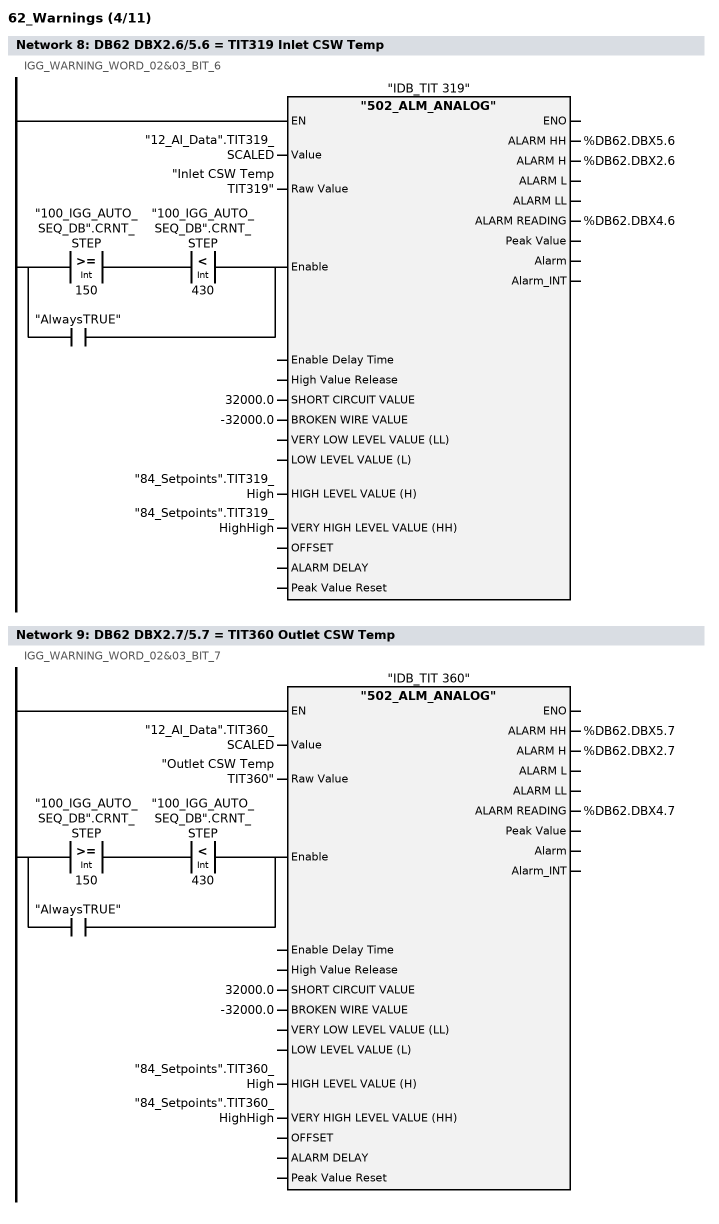
   RUNG wire#powerrail
      "IDB_TIT 319"(Enable := wire#w1, Value := "12_AI_Data".TIT319_SCALED, "Raw Value" := "Inlet CSW Temp TIT319", "SHORT CIRCUIT VALUE" := 32000.0, "BROKEN WIRE VALUE" := -32000.0, "VERY LOW LEVEL VALUE (LL)" :=, "LOW LEVEL VALUE (L)" :=, "HIGH LEVEL VALUE (H)" := "84_Setpoints".TIT319_High, "VERY HIGH LEVEL VALUE (HH)" := "84_Setpoints".TIT319_HighHigh, OFFSET :=, "ALARM DELAY" :=, "Peak Value Reset" :=, "ALARM HH" => %DB62.DBX5.6, "ALARM H" => %DB62.DBX2.6, "ALARM L" =>, "ALARM LL" =>, "ALARM READING" => %DB62.DBX4.6, "Peak Value" =>, Alarm =>, Alarm_INT =>, "Enable Delay Time" :=, "High Value Release" :=)
   END_RUNG
   RUNG wire#powerrail
      { S7_Templates := "SrcType := Int" } GE_Contact(in1 := "100_IGG_AUTO_SEQ_DB".CRNT_STEP, in2 := 150)
      { S7_Templates := "SrcType := Int" } LT_Contact(in1 := "100_IGG_AUTO_SEQ_DB".CRNT_STEP, in2 := 430)
   END_RUNG wire#w1
   RUNG wire#powerrail
      Contact( "AlwaysTRUE" )
   END_RUNG wire#w1
   // the same network as SCL:
   "IDB_TIT 319"(Value := "12_AI_Data".TIT319_SCALED,   // "502_ALM_ANALOG"
                 "Raw Value" := "Inlet CSW Temp TIT319",
                 Enable := (("100_IGG_AUTO_SEQ_DB".CRNT_STEP >= 150) AND ("100_IGG_AUTO_SEQ_DB".CRNT_STEP < 430)) OR "AlwaysTRUE",
                 "SHORT CIRCUIT VALUE" := 32000.0,
                 "BROKEN WIRE VALUE" := -32000.0,
                 "HIGH LEVEL VALUE (H)" := "84_Setpoints".TIT319_High,
                 "VERY HIGH LEVEL VALUE (HH)" := "84_Setpoints".TIT319_HighHigh,
                 "ALARM HH" => %DB62.DBX5.6,
                 "ALARM H" => %DB62.DBX2.6,
                 "ALARM READING" => %DB62.DBX4.6);
END_REGION

REGION Network 9: DB62 DBX2.7/5.7 = TIT360 Outlet CSW Temp
   // IGG_WARNING_WORD_02&03_BIT_7
   RUNG wire#powerrail
      "IDB_TIT 360"(Enable := wire#w1, Value := "12_AI_Data".TIT360_SCALED, "Raw Value" := "Outlet CSW Temp TIT360", "SHORT CIRCUIT VALUE" := 32000.0, "BROKEN WIRE VALUE" := -32000.0, "VERY LOW LEVEL VALUE (LL)" :=, "LOW LEVEL VALUE (L)" :=, "HIGH LEVEL VALUE (H)" := "84_Setpoints".TIT360_High, "VERY HIGH LEVEL VALUE (HH)" := "84_Setpoints".TIT360_HighHigh, OFFSET :=, "ALARM DELAY" :=, "Peak Value Reset" :=, "ALARM HH" => %DB62.DBX5.7, "ALARM H" => %DB62.DBX2.7, "ALARM L" =>, "ALARM LL" =>, "ALARM READING" => %DB62.DBX4.7, "Peak Value" =>, Alarm =>, Alarm_INT =>, "Enable Delay Time" :=, "High Value Release" :=)
   END_RUNG
   RUNG wire#powerrail
      { S7_Templates := "SrcType := Int" } GE_Contact(in1 := "100_IGG_AUTO_SEQ_DB".CRNT_STEP, in2 := 150)
      { S7_Templates := "SrcType := Int" } LT_Contact(in1 := "100_IGG_AUTO_SEQ_DB".CRNT_STEP, in2 := 430)
   END_RUNG wire#w1
   RUNG wire#powerrail
      Contact( "AlwaysTRUE" )
   END_RUNG wire#w1
   // the same network as SCL:
   "IDB_TIT 360"(Value := "12_AI_Data".TIT360_SCALED,   // "502_ALM_ANALOG"
                 "Raw Value" := "Outlet CSW Temp TIT360",
                 Enable := (("100_IGG_AUTO_SEQ_DB".CRNT_STEP >= 150) AND ("100_IGG_AUTO_SEQ_DB".CRNT_STEP < 430)) OR "AlwaysTRUE",
                 "SHORT CIRCUIT VALUE" := 32000.0,
                 "BROKEN WIRE VALUE" := -32000.0,
                 "HIGH LEVEL VALUE (H)" := "84_Setpoints".TIT360_High,
                 "VERY HIGH LEVEL VALUE (HH)" := "84_Setpoints".TIT360_HighHigh,
                 "ALARM HH" => %DB62.DBX5.7,
                 "ALARM H" => %DB62.DBX2.7,
                 "ALARM READING" => %DB62.DBX4.7);
END_REGION

REGION Network 10: DB62 DBX3.0/3.1/6.0/6.1 = PIT359 Inlet CSW Pressure
   // IGG_WARNING_WORD_02&04
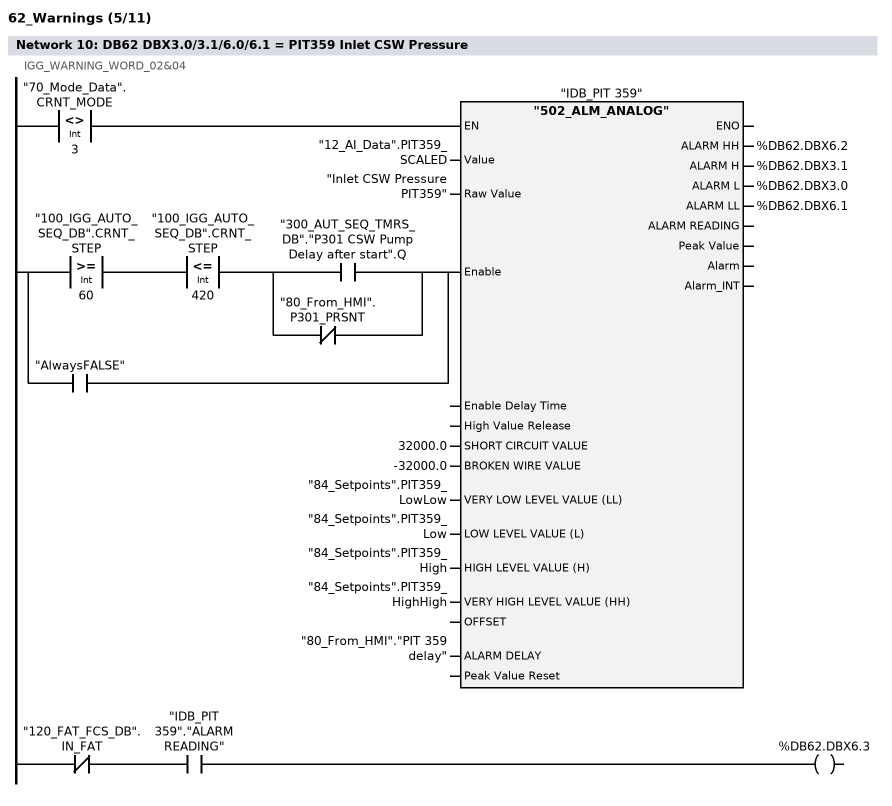
   RUNG wire#powerrail
      { S7_Templates := "SrcType := Int" } NE_Contact(in1 := "70_Mode_Data".CRNT_MODE, in2 := 3)
      "IDB_PIT 359"(Enable := wire#w2, Value := "12_AI_Data".PIT359_SCALED, "Raw Value" := "Inlet CSW Pressure PIT359", "SHORT CIRCUIT VALUE" := 32000.0, "BROKEN WIRE VALUE" := -32000.0, "VERY LOW LEVEL VALUE (LL)" := "84_Setpoints".PIT359_LowLow, "LOW LEVEL VALUE (L)" := "84_Setpoints".PIT359_Low, "HIGH LEVEL VALUE (H)" := "84_Setpoints".PIT359_High, "VERY HIGH LEVEL VALUE (HH)" := "84_Setpoints".PIT359_HighHigh, OFFSET :=, "ALARM DELAY" := "80_From_HMI"."PIT 359 delay", "Peak Value Reset" :=, "ALARM HH" => %DB62.DBX6.2, "ALARM H" => %DB62.DBX3.1, "ALARM L" => %DB62.DBX3.0, "ALARM LL" => %DB62.DBX6.1, "ALARM READING" =>, "Peak Value" =>, Alarm =>, Alarm_INT =>, "Enable Delay Time" :=, "High Value Release" :=)
   END_RUNG
   RUNG wire#powerrail
      { S7_Templates := "SrcType := Int" } GE_Contact(in1 := "100_IGG_AUTO_SEQ_DB".CRNT_STEP, in2 := 60)
      { S7_Templates := "SrcType := Int" } LE_Contact(in1 := "100_IGG_AUTO_SEQ_DB".CRNT_STEP, in2 := 420)
      wire#w1
      Contact( "300_AUT_SEQ_TMRS_DB"."P301 CSW Pump Delay after start".Q )
   END_RUNG wire#w2
   RUNG wire#w1
      I_Contact( "80_From_HMI".P301_PRSNT )
   END_RUNG wire#w2
   RUNG wire#powerrail
      Contact( "AlwaysFALSE" )
   END_RUNG wire#w2
   RUNG wire#powerrail
      I_Contact( "120_FAT_FCS_DB".IN_FAT )
      Contact( "IDB_PIT 359"."ALARM READING" )
      Coil( %DB62.DBX6.3 )
   END_RUNG
   // the same network as SCL:
   IF "70_Mode_Data".CRNT_MODE <> 3 THEN
       "IDB_PIT 359"(Value := "12_AI_Data".PIT359_SCALED,   // "502_ALM_ANALOG"
                     "Raw Value" := "Inlet CSW Pressure PIT359",
                     Enable := (("100_IGG_AUTO_SEQ_DB".CRNT_STEP >= 60) AND ("100_IGG_AUTO_SEQ_DB".CRNT_STEP <= 420) AND ("300_AUT_SEQ_TMRS_DB"."P301 CSW Pump Delay after start".Q OR NOT "80_From_HMI".P301_PRSNT)) OR "AlwaysFALSE",
                     "SHORT CIRCUIT VALUE" := 32000.0,
                     "BROKEN WIRE VALUE" := -32000.0,
                     "VERY LOW LEVEL VALUE (LL)" := "84_Setpoints".PIT359_LowLow,
                     "LOW LEVEL VALUE (L)" := "84_Setpoints".PIT359_Low,
                     "HIGH LEVEL VALUE (H)" := "84_Setpoints".PIT359_High,
                     "VERY HIGH LEVEL VALUE (HH)" := "84_Setpoints".PIT359_HighHigh,
                     "ALARM DELAY" := "80_From_HMI"."PIT 359 delay",
                     "ALARM HH" => %DB62.DBX6.2,
                     "ALARM H" => %DB62.DBX3.1,
                     "ALARM L" => %DB62.DBX3.0,
                     "ALARM LL" => %DB62.DBX6.1);
   END_IF;
   %DB62.DBX6.3 := NOT "120_FAT_FCS_DB".IN_FAT AND "IDB_PIT 359"."ALARM READING";
END_REGION

REGION Network 11: DB62 DBX3.2/3.3/3.4/3.5 = PIT316 Outlet CSW Pressure
   // IGG_WARNING_WORD_02_BIT_10&11&12&13
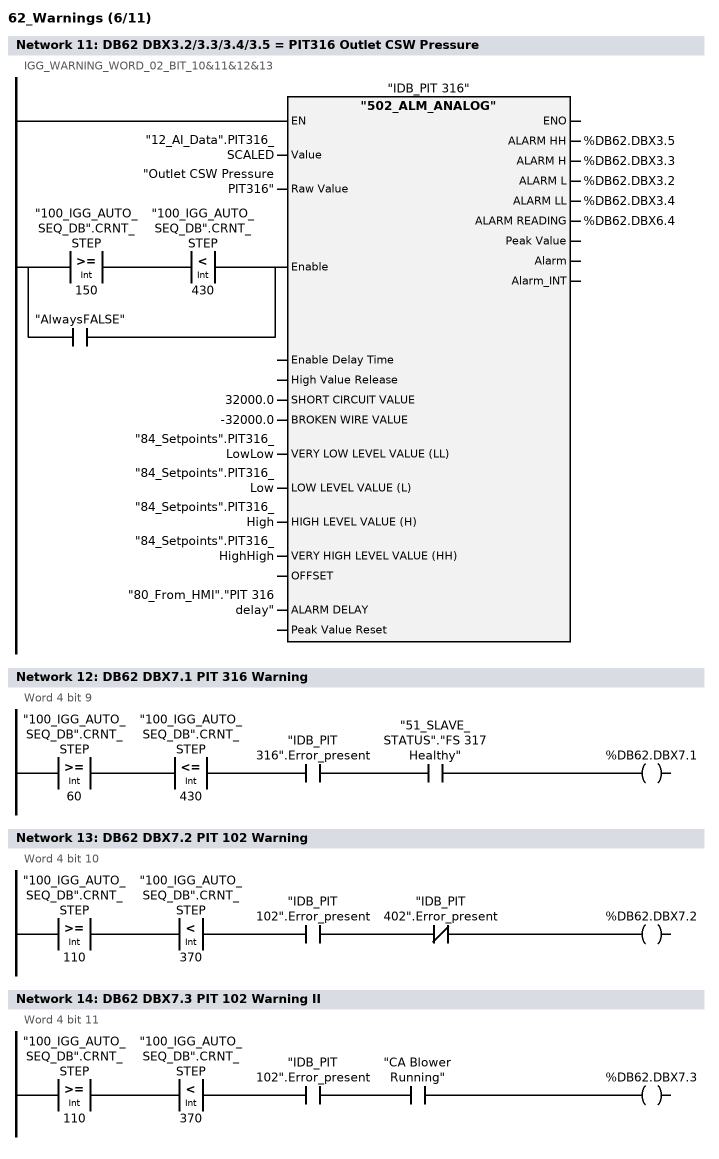
   RUNG wire#powerrail
      "IDB_PIT 316"(Enable := wire#w1, Value := "12_AI_Data".PIT316_SCALED, "Raw Value" := "Outlet CSW Pressure PIT316", "SHORT CIRCUIT VALUE" := 32000.0, "BROKEN WIRE VALUE" := -32000.0, "VERY LOW LEVEL VALUE (LL)" := "84_Setpoints".PIT316_LowLow, "LOW LEVEL VALUE (L)" := "84_Setpoints".PIT316_Low, "HIGH LEVEL VALUE (H)" := "84_Setpoints".PIT316_High, "VERY HIGH LEVEL VALUE (HH)" := "84_Setpoints".PIT316_HighHigh, OFFSET :=, "ALARM DELAY" := "80_From_HMI"."PIT 316 delay", "Peak Value Reset" :=, "ALARM HH" => %DB62.DBX3.5, "ALARM H" => %DB62.DBX3.3, "ALARM L" => %DB62.DBX3.2, "ALARM LL" => %DB62.DBX3.4, "ALARM READING" => %DB62.DBX6.4, "Peak Value" =>, Alarm =>, Alarm_INT =>, "Enable Delay Time" :=, "High Value Release" :=)
   END_RUNG
   RUNG wire#powerrail
      { S7_Templates := "SrcType := Int" } GE_Contact(in1 := "100_IGG_AUTO_SEQ_DB".CRNT_STEP, in2 := 150)
      { S7_Templates := "SrcType := Int" } LT_Contact(in1 := "100_IGG_AUTO_SEQ_DB".CRNT_STEP, in2 := 430)
   END_RUNG wire#w1
   RUNG wire#powerrail
      Contact( "AlwaysFALSE" )
   END_RUNG wire#w1
   // the same network as SCL:
   "IDB_PIT 316"(Value := "12_AI_Data".PIT316_SCALED,   // "502_ALM_ANALOG"
                 "Raw Value" := "Outlet CSW Pressure PIT316",
                 Enable := (("100_IGG_AUTO_SEQ_DB".CRNT_STEP >= 150) AND ("100_IGG_AUTO_SEQ_DB".CRNT_STEP < 430)) OR "AlwaysFALSE",
                 "SHORT CIRCUIT VALUE" := 32000.0,
                 "BROKEN WIRE VALUE" := -32000.0,
                 "VERY LOW LEVEL VALUE (LL)" := "84_Setpoints".PIT316_LowLow,
                 "LOW LEVEL VALUE (L)" := "84_Setpoints".PIT316_Low,
                 "HIGH LEVEL VALUE (H)" := "84_Setpoints".PIT316_High,
                 "VERY HIGH LEVEL VALUE (HH)" := "84_Setpoints".PIT316_HighHigh,
                 "ALARM DELAY" := "80_From_HMI"."PIT 316 delay",
                 "ALARM HH" => %DB62.DBX3.5,
                 "ALARM H" => %DB62.DBX3.3,
                 "ALARM L" => %DB62.DBX3.2,
                 "ALARM LL" => %DB62.DBX3.4,
                 "ALARM READING" => %DB62.DBX6.4);
END_REGION

REGION Network 12: DB62 DBX7.1 PIT 316 Warning
   // Word 4 bit 9
   RUNG wire#powerrail
      { S7_Templates := "SrcType := Int" } GE_Contact(in1 := "100_IGG_AUTO_SEQ_DB".CRNT_STEP, in2 := 60)
      { S7_Templates := "SrcType := Int" } LE_Contact(in1 := "100_IGG_AUTO_SEQ_DB".CRNT_STEP, in2 := 430)
      Contact( "IDB_PIT 316".Error_present )
      Contact( "51_SLAVE_STATUS"."FS 317 Healthy" )
      Coil( %DB62.DBX7.1 )
   END_RUNG
   // the same network as SCL:
   %DB62.DBX7.1 := ("100_IGG_AUTO_SEQ_DB".CRNT_STEP >= 60) AND ("100_IGG_AUTO_SEQ_DB".CRNT_STEP <= 430) AND "IDB_PIT 316".Error_present AND "51_SLAVE_STATUS"."FS 317 Healthy";
END_REGION

REGION Network 13: DB62 DBX7.2 PIT 102 Warning
   // Word 4 bit 10
   RUNG wire#powerrail
      { S7_Templates := "SrcType := Int" } GE_Contact(in1 := "100_IGG_AUTO_SEQ_DB".CRNT_STEP, in2 := 110)
      { S7_Templates := "SrcType := Int" } LT_Contact(in1 := "100_IGG_AUTO_SEQ_DB".CRNT_STEP, in2 := 370)
      Contact( "IDB_PIT 102".Error_present )
      I_Contact( "IDB_PIT 402".Error_present )
      Coil( %DB62.DBX7.2 )
   END_RUNG
   // the same network as SCL:
   %DB62.DBX7.2 := ("100_IGG_AUTO_SEQ_DB".CRNT_STEP >= 110) AND ("100_IGG_AUTO_SEQ_DB".CRNT_STEP < 370) AND "IDB_PIT 102".Error_present AND NOT "IDB_PIT 402".Error_present;
END_REGION

REGION Network 14: DB62 DBX7.3 PIT 102 Warning II
   // Word 4 bit 11
   RUNG wire#powerrail
      { S7_Templates := "SrcType := Int" } GE_Contact(in1 := "100_IGG_AUTO_SEQ_DB".CRNT_STEP, in2 := 110)
      { S7_Templates := "SrcType := Int" } LT_Contact(in1 := "100_IGG_AUTO_SEQ_DB".CRNT_STEP, in2 := 370)
      Contact( "IDB_PIT 102".Error_present )
      Contact( "CA Blower Running" )
      Coil( %DB62.DBX7.3 )
   END_RUNG
   // the same network as SCL:
   %DB62.DBX7.3 := ("100_IGG_AUTO_SEQ_DB".CRNT_STEP >= 110) AND ("100_IGG_AUTO_SEQ_DB".CRNT_STEP < 370) AND "IDB_PIT 102".Error_present AND "CA Blower Running";
END_REGION

REGION Network 15: DB62 DBX7.4 TIT 401 Warning
   // Word 4 bit 12
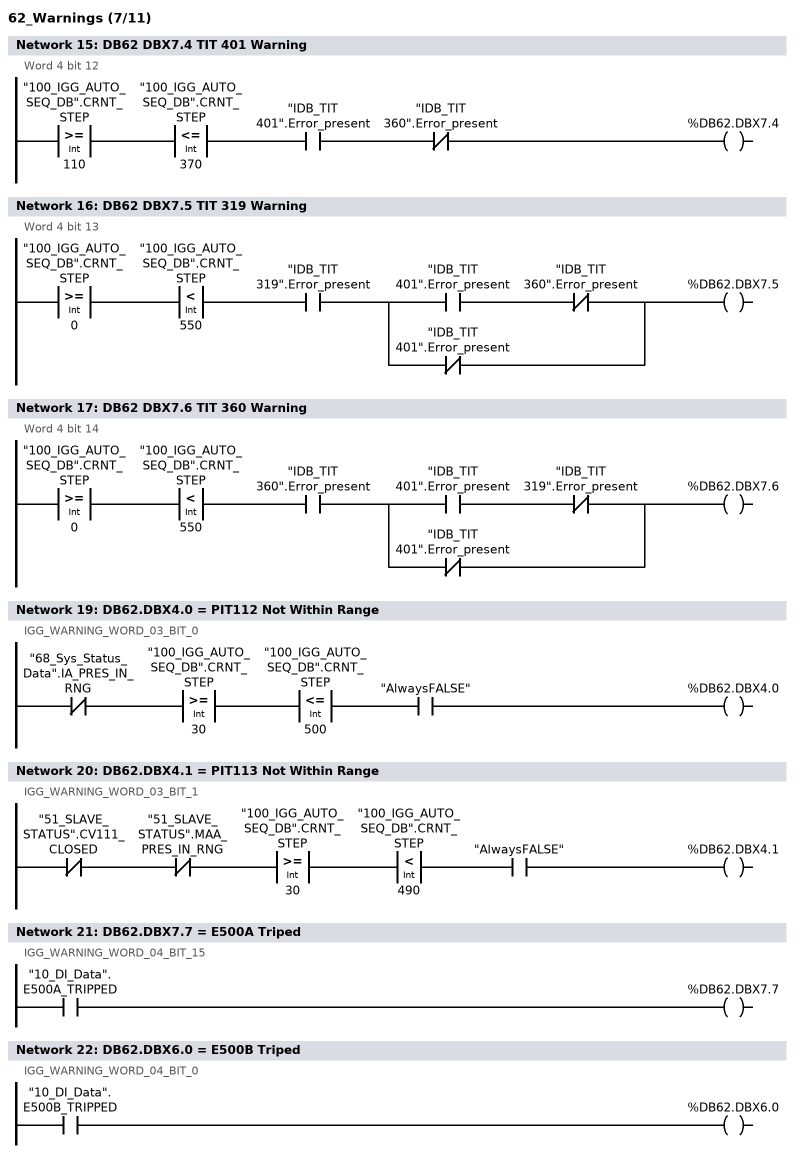
   RUNG wire#powerrail
      { S7_Templates := "SrcType := Int" } GE_Contact(in1 := "100_IGG_AUTO_SEQ_DB".CRNT_STEP, in2 := 110)
      { S7_Templates := "SrcType := Int" } LE_Contact(in1 := "100_IGG_AUTO_SEQ_DB".CRNT_STEP, in2 := 370)
      Contact( "IDB_TIT 401".Error_present )
      I_Contact( "IDB_TIT 360".Error_present )
      Coil( %DB62.DBX7.4 )
   END_RUNG
   // the same network as SCL:
   %DB62.DBX7.4 := ("100_IGG_AUTO_SEQ_DB".CRNT_STEP >= 110) AND ("100_IGG_AUTO_SEQ_DB".CRNT_STEP <= 370) AND "IDB_TIT 401".Error_present AND NOT "IDB_TIT 360".Error_present;
END_REGION

REGION Network 16: DB62 DBX7.5 TIT 319 Warning
   // Word 4 bit 13
   RUNG wire#powerrail
      { S7_Templates := "SrcType := Int" } GE_Contact(in1 := "100_IGG_AUTO_SEQ_DB".CRNT_STEP, in2 := 0)
      { S7_Templates := "SrcType := Int" } LT_Contact(in1 := "100_IGG_AUTO_SEQ_DB".CRNT_STEP, in2 := 550)
      Contact( "IDB_TIT 319".Error_present )
      wire#w1
      Contact( "IDB_TIT 401".Error_present )
      I_Contact( "IDB_TIT 360".Error_present )
      wire#w2
      Coil( %DB62.DBX7.5 )
   END_RUNG
   RUNG wire#w1
      I_Contact( "IDB_TIT 401".Error_present )
   END_RUNG wire#w2
   // the same network as SCL:
   %DB62.DBX7.5 := ("100_IGG_AUTO_SEQ_DB".CRNT_STEP >= 0) AND ("100_IGG_AUTO_SEQ_DB".CRNT_STEP < 550) AND "IDB_TIT 319".Error_present AND (("IDB_TIT 401".Error_present AND NOT "IDB_TIT 360".Error_present) OR NOT "IDB_TIT 401".Error_present);
END_REGION

REGION Network 17: DB62 DBX7.6 TIT 360 Warning
   // Word 4 bit 14
   RUNG wire#powerrail
      { S7_Templates := "SrcType := Int" } GE_Contact(in1 := "100_IGG_AUTO_SEQ_DB".CRNT_STEP, in2 := 0)
      { S7_Templates := "SrcType := Int" } LT_Contact(in1 := "100_IGG_AUTO_SEQ_DB".CRNT_STEP, in2 := 550)
      Contact( "IDB_TIT 360".Error_present )
      wire#w1
      Contact( "IDB_TIT 401".Error_present )
      I_Contact( "IDB_TIT 319".Error_present )
      wire#w2
      Coil( %DB62.DBX7.6 )
   END_RUNG
   RUNG wire#w1
      I_Contact( "IDB_TIT 401".Error_present )
   END_RUNG wire#w2
   // the same network as SCL:
   %DB62.DBX7.6 := ("100_IGG_AUTO_SEQ_DB".CRNT_STEP >= 0) AND ("100_IGG_AUTO_SEQ_DB".CRNT_STEP < 550) AND "IDB_TIT 360".Error_present AND (("IDB_TIT 401".Error_present AND NOT "IDB_TIT 319".Error_present) OR NOT "IDB_TIT 401".Error_present);
END_REGION

REGION Network 19: DB62.DBX4.0 = PIT112 Not Within Range
   // IGG_WARNING_WORD_03_BIT_0
   RUNG wire#powerrail
      I_Contact( "68_Sys_Status_Data".IA_PRES_IN_RNG )
      { S7_Templates := "SrcType := Int" } GE_Contact(in1 := "100_IGG_AUTO_SEQ_DB".CRNT_STEP, in2 := 30)
      { S7_Templates := "SrcType := Int" } LE_Contact(in1 := "100_IGG_AUTO_SEQ_DB".CRNT_STEP, in2 := 500)
      Contact( "AlwaysFALSE" )
      Coil( %DB62.DBX4.0 )
   END_RUNG
   // the same network as SCL:
   %DB62.DBX4.0 := NOT "68_Sys_Status_Data".IA_PRES_IN_RNG AND ("100_IGG_AUTO_SEQ_DB".CRNT_STEP >= 30) AND ("100_IGG_AUTO_SEQ_DB".CRNT_STEP <= 500) AND "AlwaysFALSE";
END_REGION

REGION Network 20: DB62.DBX4.1 = PIT113 Not Within Range
   // IGG_WARNING_WORD_03_BIT_1
   RUNG wire#powerrail
      I_Contact( "51_SLAVE_STATUS".CV111_CLOSED )
      I_Contact( "51_SLAVE_STATUS".MAA_PRES_IN_RNG )
      { S7_Templates := "SrcType := Int" } GE_Contact(in1 := "100_IGG_AUTO_SEQ_DB".CRNT_STEP, in2 := 30)
      { S7_Templates := "SrcType := Int" } LT_Contact(in1 := "100_IGG_AUTO_SEQ_DB".CRNT_STEP, in2 := 490)
      Contact( "AlwaysFALSE" )
      Coil( %DB62.DBX4.1 )
   END_RUNG
   // the same network as SCL:
   %DB62.DBX4.1 := NOT "51_SLAVE_STATUS".CV111_CLOSED AND NOT "51_SLAVE_STATUS".MAA_PRES_IN_RNG AND ("100_IGG_AUTO_SEQ_DB".CRNT_STEP >= 30) AND ("100_IGG_AUTO_SEQ_DB".CRNT_STEP < 490) AND "AlwaysFALSE";
END_REGION

REGION Network 21: DB62.DBX7.7 = E500A Triped
   // IGG_WARNING_WORD_04_BIT_15
   RUNG wire#powerrail
      Contact( "10_DI_Data".E500A_TRIPPED )
      Coil( %DB62.DBX7.7 )
   END_RUNG
   // the same network as SCL:
   %DB62.DBX7.7 := "10_DI_Data".E500A_TRIPPED;
END_REGION

REGION Network 22: DB62.DBX6.0 = E500B Triped
   // IGG_WARNING_WORD_04_BIT_0
   RUNG wire#powerrail
      Contact( "10_DI_Data".E500B_TRIPPED )
      Coil( %DB62.DBX6.0 )
   END_RUNG
   // the same network as SCL:
   %DB62.DBX6.0 := "10_DI_Data".E500B_TRIPPED;
END_REGION

REGION Network 23: DB62.DBX8.0 = BC PLC Power Healthy
   // IGG_WARNING_WORD_05_BIT_0
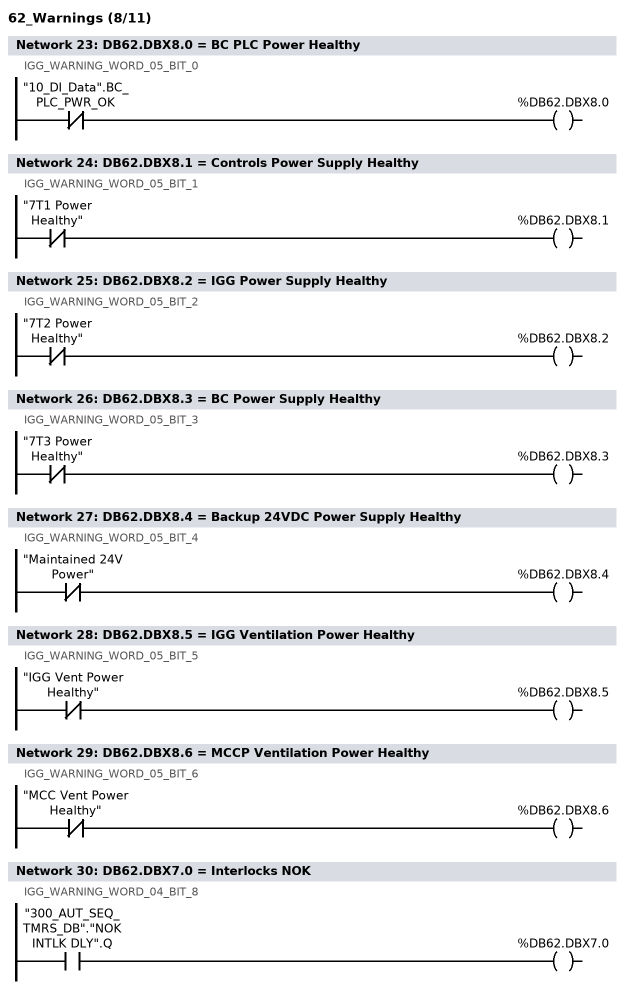
   RUNG wire#powerrail
      I_Contact( "10_DI_Data".BC_PLC_PWR_OK )
      Coil( %DB62.DBX8.0 )
   END_RUNG
   // the same network as SCL:
   %DB62.DBX8.0 := NOT "10_DI_Data".BC_PLC_PWR_OK;
END_REGION

REGION Network 24: DB62.DBX8.1 = Controls Power Supply Healthy
   // IGG_WARNING_WORD_05_BIT_1
   RUNG wire#powerrail
      I_Contact( "7T1 Power Healthy" )
      Coil( %DB62.DBX8.1 )
   END_RUNG
   // the same network as SCL:
   %DB62.DBX8.1 := NOT "7T1 Power Healthy";
END_REGION

REGION Network 25: DB62.DBX8.2 = IGG Power Supply Healthy
   // IGG_WARNING_WORD_05_BIT_2
   RUNG wire#powerrail
      I_Contact( "7T2 Power Healthy" )
      Coil( %DB62.DBX8.2 )
   END_RUNG
   // the same network as SCL:
   %DB62.DBX8.2 := NOT "7T2 Power Healthy";
END_REGION

REGION Network 26: DB62.DBX8.3 = BC Power Supply Healthy
   // IGG_WARNING_WORD_05_BIT_3
   RUNG wire#powerrail
      I_Contact( "7T3 Power Healthy" )
      Coil( %DB62.DBX8.3 )
   END_RUNG
   // the same network as SCL:
   %DB62.DBX8.3 := NOT "7T3 Power Healthy";
END_REGION

REGION Network 27: DB62.DBX8.4 = Backup 24VDC Power Supply Healthy
   // IGG_WARNING_WORD_05_BIT_4
   RUNG wire#powerrail
      I_Contact( "Maintained 24V Power" )
      Coil( %DB62.DBX8.4 )
   END_RUNG
   // the same network as SCL:
   %DB62.DBX8.4 := NOT "Maintained 24V Power";
END_REGION

REGION Network 28: DB62.DBX8.5 = IGG Ventilation Power Healthy
   // IGG_WARNING_WORD_05_BIT_5
   RUNG wire#powerrail
      I_Contact( "IGG Vent Power Healthy" )
      Coil( %DB62.DBX8.5 )
   END_RUNG
   // the same network as SCL:
   %DB62.DBX8.5 := NOT "IGG Vent Power Healthy";
END_REGION

REGION Network 29: DB62.DBX8.6 = MCCP Ventilation Power Healthy
   // IGG_WARNING_WORD_05_BIT_6
   RUNG wire#powerrail
      I_Contact( "MCC Vent Power Healthy" )
      Coil( %DB62.DBX8.6 )
   END_RUNG
   // the same network as SCL:
   %DB62.DBX8.6 := NOT "MCC Vent Power Healthy";
END_REGION

REGION Network 30: DB62.DBX7.0 = Interlocks NOK
   // IGG_WARNING_WORD_04_BIT_8
   RUNG wire#powerrail
      Contact( "300_AUT_SEQ_TMRS_DB"."NOK INTLK DLY".Q )
      Coil( %DB62.DBX7.0 )
   END_RUNG
   // the same network as SCL:
   %DB62.DBX7.0 := "300_AUT_SEQ_TMRS_DB"."NOK INTLK DLY".Q;
END_REGION

REGION Network 31: DB62.DBX9.0 = IGG HMI HeartBeat Missing
   // IGG_WARNING_WORD_05_BIT_8
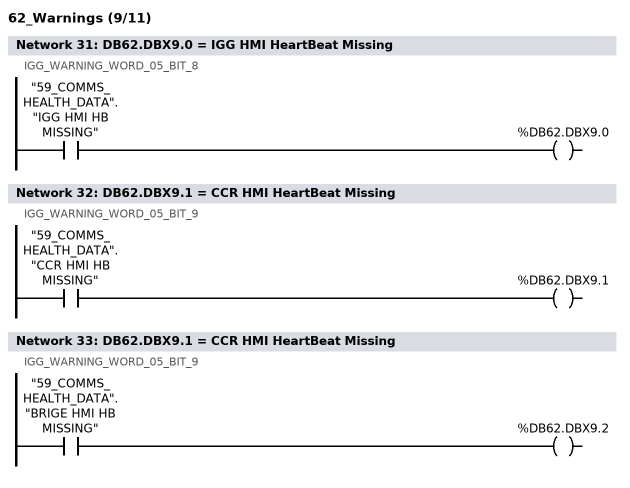
   RUNG wire#powerrail
      Contact( "59_COMMS_HEALTH_DATA"."IGG HMI HB MISSING" )
      Coil( %DB62.DBX9.0 )
   END_RUNG
   // the same network as SCL:
   %DB62.DBX9.0 := "59_COMMS_HEALTH_DATA"."IGG HMI HB MISSING";
END_REGION

REGION Network 32: DB62.DBX9.1 = CCR HMI HeartBeat Missing
   // IGG_WARNING_WORD_05_BIT_9
   RUNG wire#powerrail
      Contact( "59_COMMS_HEALTH_DATA"."CCR HMI HB MISSING" )
      Coil( %DB62.DBX9.1 )
   END_RUNG
   // the same network as SCL:
   %DB62.DBX9.1 := "59_COMMS_HEALTH_DATA"."CCR HMI HB MISSING";
END_REGION

REGION Network 33: DB62.DBX9.1 = CCR HMI HeartBeat Missing
   // IGG_WARNING_WORD_05_BIT_9
   RUNG wire#powerrail
      Contact( "59_COMMS_HEALTH_DATA"."BRIGE HMI HB MISSING" )
      Coil( %DB62.DBX9.2 )
   END_RUNG
   // the same network as SCL:
   %DB62.DBX9.2 := "59_COMMS_HEALTH_DATA"."BRIGE HMI HB MISSING";
END_REGION

REGION Network 34: Warning present
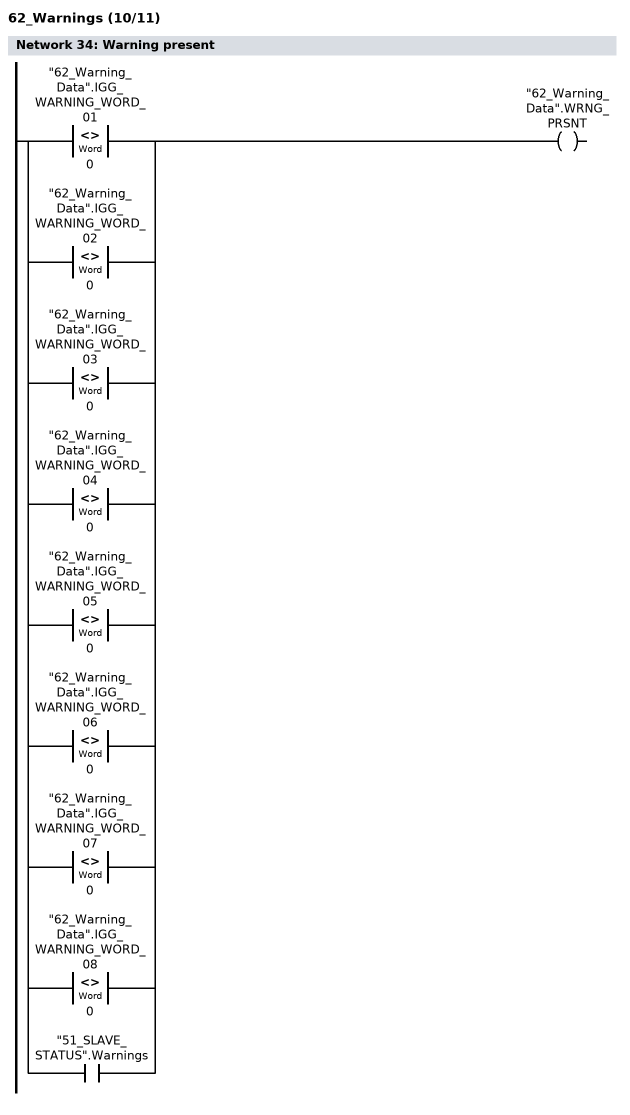
   RUNG wire#powerrail
      { S7_Templates := "SrcType := Word" } NE_Contact(in1 := "62_Warning_Data".IGG_WARNING_WORD_01, in2 := 0)
      wire#w1
      Coil( "62_Warning_Data".WRNG_PRSNT )
   END_RUNG
   RUNG wire#powerrail
      { S7_Templates := "SrcType := Word" } NE_Contact(in1 := "62_Warning_Data".IGG_WARNING_WORD_02, in2 := 0)
   END_RUNG wire#w1
   RUNG wire#powerrail
      { S7_Templates := "SrcType := Word" } NE_Contact(in1 := "62_Warning_Data".IGG_WARNING_WORD_03, in2 := 0)
   END_RUNG wire#w1
   RUNG wire#powerrail
      { S7_Templates := "SrcType := Word" } NE_Contact(in1 := "62_Warning_Data".IGG_WARNING_WORD_04, in2 := 0)
   END_RUNG wire#w1
   RUNG wire#powerrail
      { S7_Templates := "SrcType := Word" } NE_Contact(in1 := "62_Warning_Data".IGG_WARNING_WORD_05, in2 := 0)
   END_RUNG wire#w1
   RUNG wire#powerrail
      { S7_Templates := "SrcType := Word" } NE_Contact(in1 := "62_Warning_Data".IGG_WARNING_WORD_06, in2 := 0)
   END_RUNG wire#w1
   RUNG wire#powerrail
      { S7_Templates := "SrcType := Word" } NE_Contact(in1 := "62_Warning_Data".IGG_WARNING_WORD_07, in2 := 0)
   END_RUNG wire#w1
   RUNG wire#powerrail
      { S7_Templates := "SrcType := Word" } NE_Contact(in1 := "62_Warning_Data".IGG_WARNING_WORD_08, in2 := 0)
   END_RUNG wire#w1
   RUNG wire#powerrail
      Contact( "51_SLAVE_STATUS".Warnings )
   END_RUNG wire#w1
   // the same network as SCL:
   "62_Warning_Data".WRNG_PRSNT := ("62_Warning_Data".IGG_WARNING_WORD_01 <> 0) OR ("62_Warning_Data".IGG_WARNING_WORD_02 <> 0) OR ("62_Warning_Data".IGG_WARNING_WORD_03 <> 0) OR ("62_Warning_Data".IGG_WARNING_WORD_04 <> 0) OR ("62_Warning_Data".IGG_WARNING_WORD_05 <> 0) OR ("62_Warning_Data".IGG_WARNING_WORD_06 <> 0) OR ("62_Warning_Data".IGG_WARNING_WORD_07 <> 0) OR ("62_Warning_Data".IGG_WARNING_WORD_08 <> 0) OR "51_SLAVE_STATUS".Warnings;
END_REGION

REGION Network 35: New Warning Check
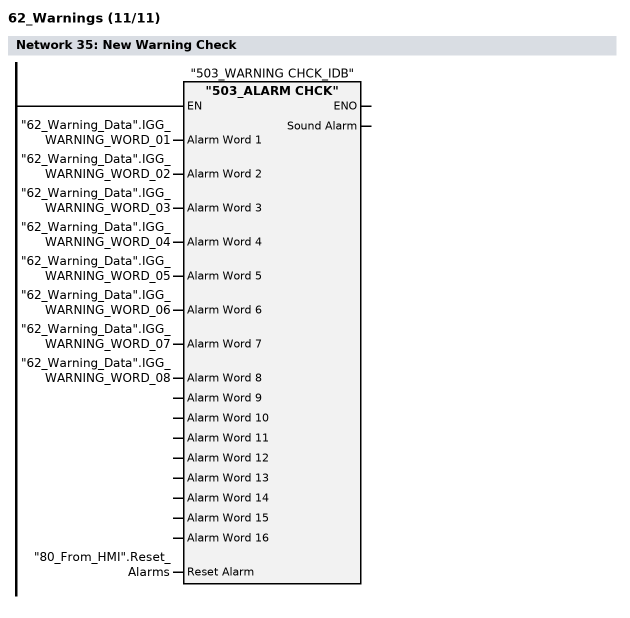
   RUNG wire#powerrail
      "503_WARNING CHCK_IDB"("Alarm Word 1" := "62_Warning_Data".IGG_WARNING_WORD_01, "Alarm Word 2" := "62_Warning_Data".IGG_WARNING_WORD_02, "Alarm Word 3" := "62_Warning_Data".IGG_WARNING_WORD_03, "Alarm Word 4" := "62_Warning_Data".IGG_WARNING_WORD_04, "Alarm Word 5" := "62_Warning_Data".IGG_WARNING_WORD_05, "Alarm Word 6" := "62_Warning_Data".IGG_WARNING_WORD_06, "Alarm Word 7" := "62_Warning_Data".IGG_WARNING_WORD_07, "Alarm Word 8" := "62_Warning_Data".IGG_WARNING_WORD_08, "Alarm Word 9" :=, "Alarm Word 10" :=, "Alarm Word 11" :=, "Alarm Word 12" :=, "Alarm Word 13" :=, "Alarm Word 14" :=, "Alarm Word 15" :=, "Alarm Word 16" :=, "Reset Alarm" := "80_From_HMI".Reset_Alarms, "Sound Alarm" =>)
   END_RUNG
   // the same network as SCL:
   "503_WARNING CHCK_IDB"("Alarm Word 1" := "62_Warning_Data".IGG_WARNING_WORD_01,   // "503_ALARM CHCK"
                          "Alarm Word 2" := "62_Warning_Data".IGG_WARNING_WORD_02,
                          "Alarm Word 3" := "62_Warning_Data".IGG_WARNING_WORD_03,
                          "Alarm Word 4" := "62_Warning_Data".IGG_WARNING_WORD_04,
                          "Alarm Word 5" := "62_Warning_Data".IGG_WARNING_WORD_05,
                          "Alarm Word 6" := "62_Warning_Data".IGG_WARNING_WORD_06,
                          "Alarm Word 7" := "62_Warning_Data".IGG_WARNING_WORD_07,
                          "Alarm Word 8" := "62_Warning_Data".IGG_WARNING_WORD_08,
                          "Reset Alarm" := "80_From_HMI".Reset_Alarms);
END_REGION
END_FUNCTION

FUNCTION "68_Sys_Status" : Void   // FC68, LAD
TITLE = System Status
{ S7_Optimized_Access := 'TRUE' }
AUTHOR : JRS
VERSION : 0.1
// For the determination of specific system status information as required by the code
   VAR_TEMP   // added for the SCL form of the ladder/FBD networks
      _w1 : Bool;
      _w2 : Bool;
   END_VAR
BEGIN

REGION Network 1: Valves At Initial
   // All valves in initial state
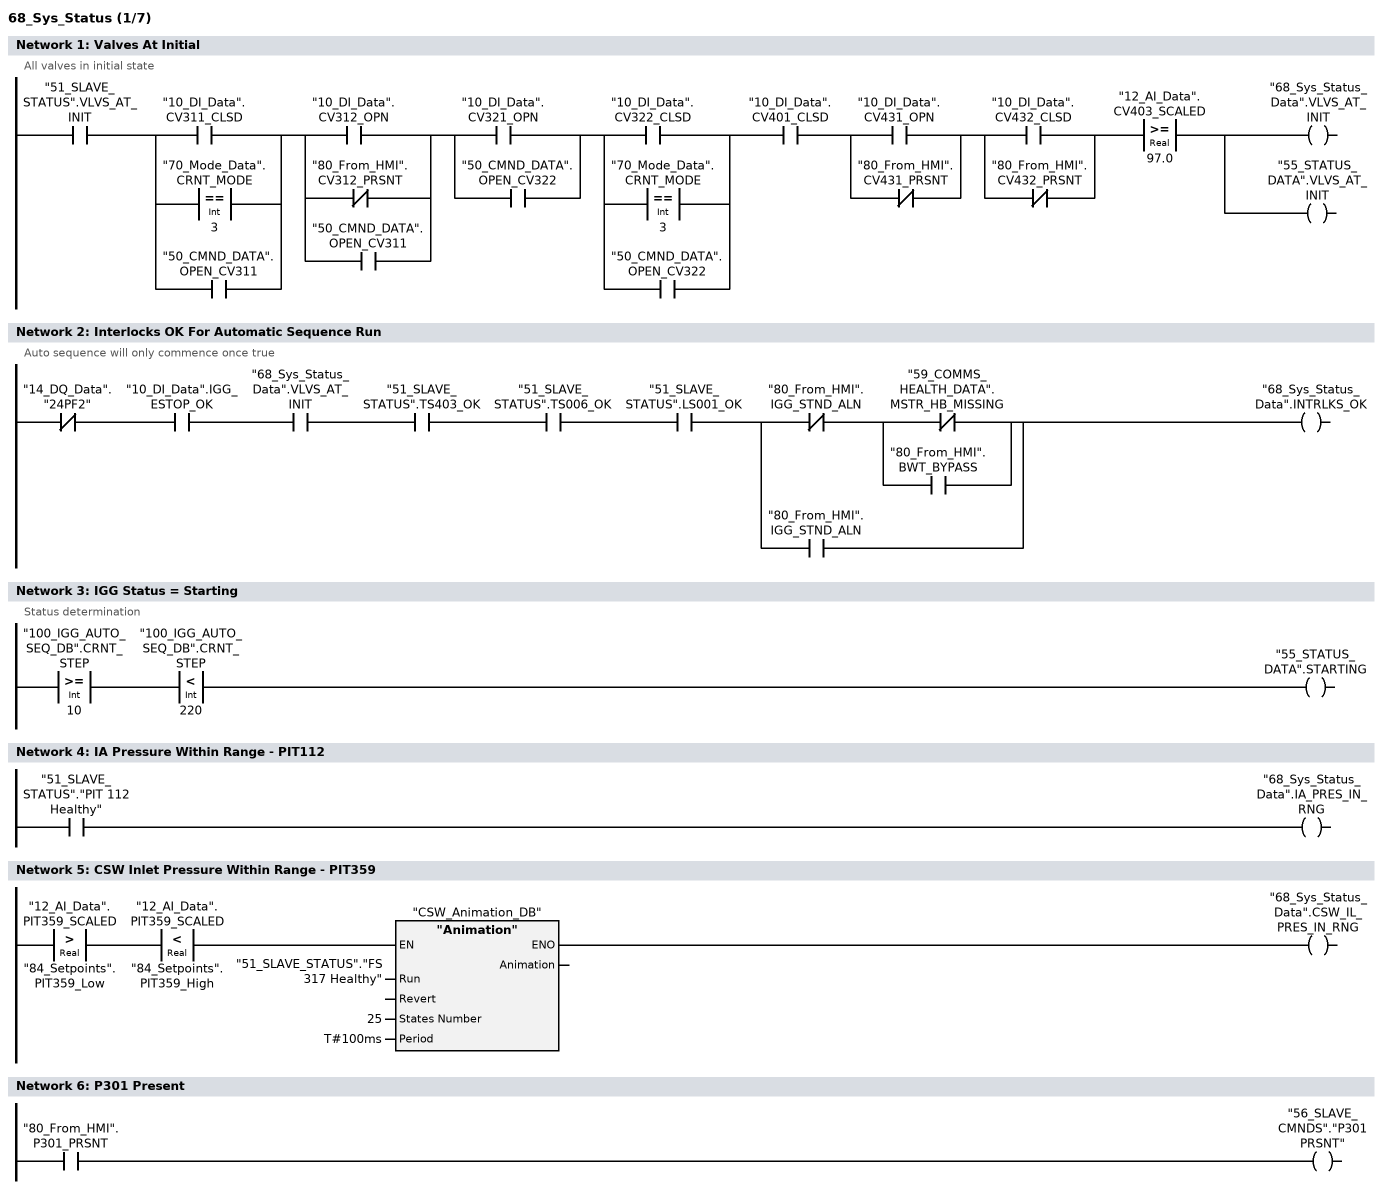
   RUNG wire#powerrail
      Contact( "51_SLAVE_STATUS".VLVS_AT_INIT )
      wire#w1
      Contact( "10_DI_Data".CV311_CLSD )
      wire#w2
      Contact( "10_DI_Data".CV312_OPN )
      wire#w3
      Contact( "10_DI_Data".CV321_OPN )
      wire#w4
      Contact( "10_DI_Data".CV322_CLSD )
      wire#w5
      Contact( "10_DI_Data".CV401_CLSD )
      wire#w6
      Contact( "10_DI_Data".CV431_OPN )
      wire#w7
      Contact( "10_DI_Data".CV432_CLSD )
      wire#w8
      { S7_Templates := "SrcType := Real" } GE_Contact(in1 := "12_AI_Data".CV403_SCALED, in2 := 97.0)
      wire#w9
      Coil( "68_Sys_Status_Data".VLVS_AT_INIT )
   END_RUNG
   RUNG wire#w1
      { S7_Templates := "SrcType := Int" } EQ_Contact(in1 := "70_Mode_Data".CRNT_MODE, in2 := 3)
   END_RUNG wire#w2
   RUNG wire#w1
      Contact( "50_CMND_DATA".OPEN_CV311 )
   END_RUNG wire#w2
   RUNG wire#w2
      I_Contact( "80_From_HMI".CV312_PRSNT )
   END_RUNG wire#w3
   RUNG wire#w2
      Contact( "50_CMND_DATA".OPEN_CV311 )
   END_RUNG wire#w3
   RUNG wire#w3
      Contact( "50_CMND_DATA".OPEN_CV322 )
   END_RUNG wire#w4
   RUNG wire#w4
      { S7_Templates := "SrcType := Int" } EQ_Contact(in1 := "70_Mode_Data".CRNT_MODE, in2 := 3)
   END_RUNG wire#w5
   RUNG wire#w4
      Contact( "50_CMND_DATA".OPEN_CV322 )
   END_RUNG wire#w5
   RUNG wire#w6
      I_Contact( "80_From_HMI".CV431_PRSNT )
   END_RUNG wire#w7
   RUNG wire#w7
      I_Contact( "80_From_HMI".CV432_PRSNT )
   END_RUNG wire#w8
   RUNG wire#w9
      Coil( "55_STATUS_DATA".VLVS_AT_INIT )
   END_RUNG
   // the same network as SCL:
   "68_Sys_Status_Data".VLVS_AT_INIT := "51_SLAVE_STATUS".VLVS_AT_INIT AND ("10_DI_Data".CV311_CLSD OR ("70_Mode_Data".CRNT_MODE = 3) OR "50_CMND_DATA".OPEN_CV311) AND ("10_DI_Data".CV312_OPN OR NOT "80_From_HMI".CV312_PRSNT OR "50_CMND_DATA".OPEN_CV311) AND ("10_DI_Data".CV321_OPN OR "50_CMND_DATA".OPEN_CV322) AND ("10_DI_Data".CV322_CLSD OR ("70_Mode_Data".CRNT_MODE = 3) OR "50_CMND_DATA".OPEN_CV322) AND "10_DI_Data".CV401_CLSD AND ("10_DI_Data".CV431_OPN OR NOT "80_From_HMI".CV431_PRSNT) AND ("10_DI_Data".CV432_CLSD OR NOT "80_From_HMI".CV432_PRSNT) AND ("12_AI_Data".CV403_SCALED >= 97.0);
   "55_STATUS_DATA".VLVS_AT_INIT := "68_Sys_Status_Data".VLVS_AT_INIT;
END_REGION

REGION Network 2: Interlocks OK For Automatic Sequence Run
   // Auto sequence will only commence once true
   RUNG wire#powerrail
      I_Contact( "14_DQ_Data"."24PF2" )
      Contact( "10_DI_Data".IGG_ESTOP_OK )
      Contact( "68_Sys_Status_Data".VLVS_AT_INIT )
      Contact( "51_SLAVE_STATUS".TS403_OK )
      Contact( "51_SLAVE_STATUS".TS006_OK )
      Contact( "51_SLAVE_STATUS".LS001_OK )
      wire#w1
      I_Contact( "80_From_HMI".IGG_STND_ALN )
      wire#w2
      I_Contact( "59_COMMS_HEALTH_DATA".MSTR_HB_MISSING )
      wire#w3
      Coil( "68_Sys_Status_Data".INTRLKS_OK )
   END_RUNG
   RUNG wire#w2
      Contact( "80_From_HMI".BWT_BYPASS )
   END_RUNG wire#w3
   RUNG wire#w1
      Contact( "80_From_HMI".IGG_STND_ALN )
   END_RUNG wire#w3
   // the same network as SCL:
   "68_Sys_Status_Data".INTRLKS_OK := NOT "14_DQ_Data"."24PF2" AND "10_DI_Data".IGG_ESTOP_OK AND "68_Sys_Status_Data".VLVS_AT_INIT AND "51_SLAVE_STATUS".TS403_OK AND "51_SLAVE_STATUS".TS006_OK AND "51_SLAVE_STATUS".LS001_OK AND ((NOT "80_From_HMI".IGG_STND_ALN AND (NOT "59_COMMS_HEALTH_DATA".MSTR_HB_MISSING OR "80_From_HMI".BWT_BYPASS)) OR "80_From_HMI".IGG_STND_ALN);
END_REGION

REGION Network 3: IGG Status = Starting
   // Status determination
   RUNG wire#powerrail
      { S7_Templates := "SrcType := Int" } GE_Contact(in1 := "100_IGG_AUTO_SEQ_DB".CRNT_STEP, in2 := 10)
      { S7_Templates := "SrcType := Int" } LT_Contact(in1 := "100_IGG_AUTO_SEQ_DB".CRNT_STEP, in2 := 220)
      Coil( "55_STATUS_DATA".STARTING )
   END_RUNG
   // the same network as SCL:
   "55_STATUS_DATA".STARTING := ("100_IGG_AUTO_SEQ_DB".CRNT_STEP >= 10) AND ("100_IGG_AUTO_SEQ_DB".CRNT_STEP < 220);
END_REGION

REGION Network 4: IA Pressure Within Range - PIT112
   RUNG wire#powerrail
      Contact( "51_SLAVE_STATUS"."PIT 112 Healthy" )
      Coil( "68_Sys_Status_Data".IA_PRES_IN_RNG )
   END_RUNG
   // the same network as SCL:
   "68_Sys_Status_Data".IA_PRES_IN_RNG := "51_SLAVE_STATUS"."PIT 112 Healthy";
END_REGION

REGION Network 5: CSW Inlet Pressure Within Range - PIT359
   RUNG wire#powerrail
      { S7_Templates := "SrcType := Real" } GT_Contact(in1 := "12_AI_Data".PIT359_SCALED, in2 := "84_Setpoints".PIT359_Low)
      { S7_Templates := "SrcType := Real" } LT_Contact(in1 := "12_AI_Data".PIT359_SCALED, in2 := "84_Setpoints".PIT359_High)
      "CSW_Animation_DB"(Run := "51_SLAVE_STATUS"."FS 317 Healthy", Revert :=, "States Number" := 25, Period := T#100ms, Animation =>)
      Coil( "68_Sys_Status_Data".CSW_IL_PRES_IN_RNG )
   END_RUNG
   // the same network as SCL:
   "CSW_Animation_DB"(EN := ("12_AI_Data".PIT359_SCALED > "84_Setpoints".PIT359_Low) AND ("12_AI_Data".PIT359_SCALED < "84_Setpoints".PIT359_High),   // "Animation"
                      Run := "51_SLAVE_STATUS"."FS 317 Healthy",
                      "States Number" := 25,
                      Period := T#100ms,
                      ENO => #_w1);
   "68_Sys_Status_Data".CSW_IL_PRES_IN_RNG := #_w1;
END_REGION

REGION Network 6: P301 Present
   RUNG wire#powerrail
      Contact( "80_From_HMI".P301_PRSNT )
      Coil( "56_SLAVE_CMNDS"."P301 PRSNT" )
   END_RUNG
   // the same network as SCL:
   "56_SLAVE_CMNDS"."P301 PRSNT" := "80_From_HMI".P301_PRSNT;
END_REGION

REGION Network 7: Fuel Pump A Runt Time - E500A
